(* Logix 5000 project; controller PLC_MCC1201_220AP1 vendor 1 type 14 code 164 rev 35.11; software revision 35.00; part 4 of 25 *)

        [201]   // Flaw Tail Lane Ptr
        [202]   // Flaw Tail Offset Ptr
        [203]   // Count at Sync Pulse to Host MSW
        [204]   // Count at Sync Pulse to Host LSW
        [205]   // Count at Data Request to Host MSW
        [206]   // Count at Data Request to Host LSW
        [207]   // Host Integer location for the number of 1 Meter Pulses(0-39)
        [208]   // Host location for 1/10 millimeter position since last 1 Meter
        [209].0   // Data Request to Host
        [209].1   // Cover Closed to Host
        [209].2   // Use Insp. Booth P.B. only, to host
        [209].4   // Cross Break in Progress to Host
        [209].6   // Image Automation in Alarm to Host
        [209].7   // Image Automation Watchdog Alarm to Host
        [210]   // Lehr Speed to Host
        [211]   // Manual Inspection Flaw Pos. MSW
        [212]   // Manual Inspection Flaw Pos. LSW
        [234]   // Time for last Meter in 0.01 sec
        [237]   // Copy of Count at Data Request to Host MSW
        [238]   // Copy of Count at Data Request to Host LSW
        [209].5   // Crush All Plates to Host
        [209].8   // Always True Signal to Host
   N44 : DINT[213] := ([0] := -1, [2] := -1, [4] := -1, [6] := -1, [8] := -1, [10] := -1, [12] := -1, [14] := -1, [16] := -1, [18] := -1, [20] := -1, [22] := -1, [24] := -1, [26] := -1, [28] := -1, [30] := -1, [32] := -1, [34] := -1, [36] := -1, [38] := -1, [40] := -1, [42] := -1, [44] := -1, [46] := -1, [48] := -1, [50] := -1, [52] := -1, [54] := -1, [56] := -1, [58] := -1, [60] := -1, [62] := -1, [64] := -1, [66] := -1, [68] := -1, [70] := -1, [72] := -1, [74] := -1, [76] := -1, [78] := -1, [80] := -1, [82] := -1, [84] := -1, [86] := -1, [88] := -1, [90] := -1, [92] := -1, [94] := -1, [96] := -1, [98] := -1, [200] := -1);
   N45 : DINT[58] := ([4] := 244, [5] := 129, [6] := 810, [21] := -21856, [23] := 1296, [24] := 253, [26] := 8192, [27] := 5376, [29] := 20480, [30] := 8192, [31] := 8192, [32] := 8192, [33] := 8192, [34] := 8192, [35] := 8192, [36] := 8192, [37] := 8192, [38] := 8192, [39] := 8192, [40] := 8192, [41] := 8192);
   N46 : DINT[7] := ([0] := 142);
        [0]   // Strain Count
        [1]   // Strain Status
        [2]   // Start Strain Cycle
        [3]   // Bar Disable For Reliance
   N47 : DINT[200] := ([0] := 296, [1] := 523, [2] := 448, [3] := 301, [4] := 248, [5] := 289, [6] := 298, [7] := 292, [8] := 287, [9] := 256, [10] := 239, [11] := 185, [12] := 175, [13] := 141, [14] := 116, [15] := 67, [16] := 50, [17] := 74, [18] := 73, [19] := 79, [20] := 75, [21] := 92, [22] := 90, [23] := 90, [24] := 73, [25] := 47, [26] := 29, [27] := 1, [28] := 36, [29] := 39, [30] := 45, [31] := 76, [32] := 75, [33] := 92, [34] := 73, [35] := 84, [36] := 96, [37] := 90, [38] := 74, [39] := 56, [40] := 68, [41] := 72, [42] := 71, [43] := 81, [44] := 78, [45] := 86, [46] := 85, [47] := 88, [48] := 96, [49] := 76, [50] := 54, [51] := 39, [52] := 68, [53] := 89, [54] := 93, [55] := 100, [56] := 103, [57] := 111, [58] := 100, [59] := 114,
        [60] := 125, [61] := 115, [62] := 111, [63] := 109, [64] := 102, [65] := 135, [66] := 135, [67] := 131, [68] := 153, [69] := 136, [70] := 126, [71] := 125, [72] := 122, [73] := 100, [74] := 84, [75] := 82, [76] := 111, [77] := 126, [78] := 127, [79] := 115, [80] := 128, [81] := 123, [82] := 138, [83] := 123, [84] := 110, [85] := 83, [86] := 62, [87] := 68, [88] := 91, [89] := 82, [90] := 100, [91] := 129, [92] := 129, [93] := 110, [94] := 118, [95] := 103, [96] := 121, [97] := 96, [98] := 94, [99] := 107, [100] := 129, [101] := 119, [102] := 123, [103] := 123, [104] := 95, [105] := 101, [106] := 90, [107] := 82, [108] := 78, [109] := 39, [110] := 37, [111] := 62, [112] := 77, [113] := 64, [114] := 68, [115] := 81, [116] := 94, [117] := 83, [118] := 94, [119] := 109,
        [120] := 118, [121] := 123, [122] := 132, [123] := 160, [124] := 190, [125] := 245, [126] := 254, [127] := 295, [128] := 313, [129] := 349, [130] := 383, [131] := 378, [132] := 331, [133] := 284, [134] := 363, [135] := 508, [136] := 87, [137] := 124, [138] := 115, [139] := 132, [140] := 122, [141] := 121, [142] := 126, [143] := 184, [144] := 171, [145] := 122, [146] := 134, [147] := 224, [148] := 143, [149] := 179, [150] := 182, [151] := 488, [152] := 583, [153] := 710, [154] := 493, [155] := 464, [156] := 456, [157] := 470, [158] := 458, [159] := 453, [160] := 458, [161] := 459, [162] := 459, [163] := 464, [164] := 470, [165] := 437, [166] := 467, [167] := 455, [168] := 446, [169] := 426, [170] := 443, [171] := 429, [172] := 422, [173] := 436, [174] := 449, [175] := 433, [176] := 452, [177] := 425, [178] := 447, [179] := 437,
        [180] := 443, [181] := 420, [182] := 440, [183] := 439, [184] := 417, [185] := 427, [186] := 428, [187] := 431, [188] := 429, [189] := 437, [190] := 437, [191] := 419, [192] := 435, [193] := 420, [194] := 421, [195] := 427, [196] := 430, [197] := 439, [198] := 423, [199] := 451);
   N48 : DINT[200] := ([0] := 1032, [1] := 1100, [2] := 1101, [3] := 1081, [4] := 1082, [5] := 1097, [6] := 1100, [7] := 1108, [8] := 1119, [9] := 1115, [10] := 1120, [11] := 1115, [12] := 1114, [13] := 1110, [14] := 1106, [15] := 1095, [16] := 1102, [17] := 1112, [18] := 1121, [19] := 1118, [20] := 1123, [21] := 1120, [22] := 1119, [23] := 1114, [24] := 1118, [25] := 1115, [26] := 1111, [27] := 1106, [28] := 1114, [29] := 1120, [30] := 1125, [31] := 1129, [32] := 1126, [33] := 1119, [34] := 1118, [35] := 1126, [36] := 1126, [37] := 1126, [38] := 1117, [39] := 1117, [40] := 1118, [41] := 1124, [42] := 1124, [43] := 1125, [44] := 1124, [45] := 1128, [46] := 1128, [47] := 1130, [48] := 1132, [49] := 1124, [50] := 1114, [51] := 1115, [52] := 1124, [53] := 1136, [54] := 1133, [55] := 1132, [56] := 1133, [57] := 1133, [58] := 1137, [59] := 1140,
        [60] := 1136, [61] := 1129, [62] := 1125, [63] := 1128, [64] := 1126, [65] := 1134, [66] := 1133, [67] := 1136, [68] := 1139, [69] := 1131, [70] := 1132, [71] := 1140, [72] := 1129, [73] := 1127, [74] := 1115, [75] := 1131, [76] := 1133, [77] := 1135, [78] := 1132, [79] := 1138, [80] := 1140, [81] := 1136, [82] := 1140, [83] := 1138, [84] := 1132, [85] := 1123, [86] := 1128, [87] := 1127, [88] := 1137, [89] := 1133, [90] := 1134, [91] := 1135, [92] := 1132, [93] := 1127, [94] := 1131, [95] := 1129, [96] := 1126, [97] := 1117, [98] := 1120, [99] := 1134, [100] := 1129, [101] := 1130, [102] := 1130, [103] := 1121, [104] := 1119, [105] := 1115, [106] := 1115, [107] := 1116, [108] := 1105, [109] := 1098, [110] := 1102, [111] := 1116, [112] := 1113, [113] := 1108, [114] := 1108, [115] := 1108, [116] := 1113, [117] := 1108, [118] := 1108, [119] := 1107,
        [120] := 1097, [121] := 1094, [122] := 1097, [123] := 1094, [124] := 1092, [125] := 1091, [126] := 1093, [127] := 1089, [128] := 1084, [129] := 1091, [130] := 1089, [131] := 1082, [132] := 1065, [133] := 1068, [134] := 1099, [135] := 1083, [136] := 838, [137] := 839, [138] := 830, [139] := 832, [140] := 829, [141] := 828, [142] := 829, [143] := 827, [144] := 827, [145] := 850, [146] := 846, [147] := 842, [148] := 848, [149] := 846, [150] := 870, [151] := 1103, [152] := 1068, [153] := 1082, [154] := 1031, [155] := 1033, [156] := 1029, [157] := 1034, [158] := 1034, [159] := 1033, [160] := 1035, [161] := 1039, [162] := 1040, [163] := 1038, [164] := 1041, [165] := 1045, [166] := 1041, [167] := 1040, [168] := 1042, [169] := 1041, [170] := 1044, [171] := 1045, [172] := 1040, [173] := 1042, [174] := 1045, [175] := 1040, [176] := 1042, [177] := 1032, [178] := 1041, [179] := 1049,
        [180] := 1042, [181] := 1046, [182] := 1045, [183] := 1043, [184] := 1044, [185] := 1048, [186] := 1047, [187] := 1043, [188] := 1048, [189] := 1040, [190] := 1040, [191] := 1043, [192] := 1041, [193] := 1038, [194] := 1041, [195] := 1042, [196] := 1039, [197] := 1044, [198] := 1038, [199] := 1042);
   N50 : DINT[40] := ([5] := 6278, [7] := 1);
        [39].0   // NO1 CRUSHER Crusher is up and in manual alarm horn has been acknowledged.
   N500 : DINT[24] := ([1] := 1755, [2] := 1755, [3] := 1755, [4] := 1755, [5] := 1755, [6] := 1755, [7] := 1755);
   N501 : DINT[25] := ([1] := 21, [2] := 21, [3] := 21, [4] := 21, [5] := 71, [6] := 71, [7] := 6);
   N502 : DINT[25] := ([1] := 361, [2] := 361, [3] := 361, [4] := 361, [5] := 361, [6] := 361, [7] := 361);
   N504 : DINT[25] := ([1] := 2975, [2] := 2975, [3] := 2975, [4] := 2975, [5] := 3600, [6] := 3600, [7] := 4398);
   N505 : DINT[25] := ([1] := 4229, [2] := 4229, [3] := 4229, [4] := 4229, [5] := 1514, [6] := 1514, [7] := 21881);
   N506 : DINT[25];
   N507 : DINT[25] := ([1] := 765, [2] := 765, [3] := 766, [4] := 766, [5] := 1493, [6] := 1493, [7] := 103, [17] := 1816, [18] := 1816, [24] := 2750);
        [17]   // SPEED CALC Current Command freq. For washer Sponges
        [24]   // SPEED CALC Current Lehr spd + 1.5% Times 10
   N53 : DINT[10];
        [0]   // Disable Y-cuts Information Written FROM Host computer
        [1]   // MANUAL INSPCTN Reject flaw Q.A. Flaw Lamps host Write word
        [2].3   // HOST WRITE Inhibit bit For Trim Deck E-stop
        [2].4   // HOST WRITE Inhibit bit For Critical Failure
        [2].5   // HOST WRITE Inhibit bit For trim Deck drive Fault
        [2].7   // HOST WRITE Inhibit bit for Mainline Backup
        [2].8   // HOST WRITE Inhibit bit for Drive system E-stop
        [2].10   // HOST WRITE Inhibit bit for Sec. Trans. Drive fault
        [2].11   // Host Critical Alarm Present
        [2].12   // View TEC15V alarm present
        [2].13   // APC Low Alarm
        [3].0   // From Host Enable 37B's REV controls
        [5].0   // ISRA 5D System QC Request Signal
        [5].1   // ISRA 5D System Cut Signal
        [8].6   // Z200 Reset Alarms
        [8]   // HOST WRITE DATA: ZONE 200 (Cutting Area) HMI Commands
        [8].0   // Z200 Start Cycle
        [8].3   // Z200 Stop Cleaning
        [8].1   // Z200 Stop Cycle
        [8].4   // Z200 Zone in Automatic
        [8].5   // Z200 Zone in Manual
        [8].2   // Z200 Start Cleaning
        [7]   // HOST WRITE DATA: ZONE UPS (Drop Conveyor Area) HMI Commands
        [7].0   // ZUPS Start Cycle
        [7].1   // ZUPS Stop Cycle
        [7].2   // ZUPS Start Cleaning
        [7].3   // ZUPS Stop Cleaning
        [7].4   // ZUPS Zone in Automatic
        [7].5   // ZUPS Zone in Manual
        [7].6   // ZUPS Reset Alarms
   N53_HOST : INT[10];
   N54 : DINT[501] := ([200] := 516, [201] := 1844, [202] := 516, [203] := 516, [204] := 516, [206] := 4, [207] := 31, [208] := 514, [211] := 176, [239] := 16, [240] := -65524, [244] := 4096, [246] := 512, [247] := 256, [248] := 512, [249] := 1, [250] := 15, [251] := 17, [252] := 12, [253] := 8, [254] := 44, [255] := 27, [256] := 15, [257] := 13, [258] := 10, [259] := 10, [260] := 481, [261] := 480, [262] := 481, [264] := -32287, [265] := 10, [266] := 110, [270] := 132, [271] := 164, [273] := 1, [274] := 1, [275] := 1, [276] := 1, [277] := 1, [281] := -32768, [341] := 133, [368] := -11667, [410] := 9, [411] := 510, [420] := 6234);
        [200].1   // RIBBON WASHER BRUSH #1 AUTO Mode Bit
        [200].2   // RIBBON WASHER BRUSH #1 MANUAL Mode Bit
        [200].3   // RIBBON WASHER BRUSH #1 ON Sw. Inputs
        [200].4   // RIBBON WASHER BRUSH #1 OFF Sw. Inputs
        [200].5   // RIBBON WASHER BRUSH #1 UPPER RETRACT Sw. Inputs
        [200].6   // RIBBON WASHER BRUSH #1 UPPER CONVERGE Sw. Inputs
        [200].7   // RIBBON WASHER BRUSH #1 LOWER RETRACT Sw. Inputs
        [200].8   // RIBBON WASHER BRUSH #1 LOWER CONVERGE Sw. Inputs
        [200].9   // RIBBON WASHER BRUSH #1 Manual Mode Lamp
        [200].10   // RIBBON WASHER BRUSH #1 OFF selected Manual mode
        [202].1   // RIBBON WASHER SPONGE UNIT AUTO Mode Bit
        [202].2   // RIBBON WASHER SPONGE UNIT MANUAL Mode Bit
        [202].3   // RIBBON WASHER SPONGE UNIT ON Sw. Inputs
        [202].4   // RIBBON WASHER SPONGE UNIT OFF Sw. Inputs
        [202].5   // RIBBON WASHER SPONGE UNIT UPPER RETRACT Sw. Inputs
        [202].6   // RIBBON WASHER SPONGE UNIT UPPER CONVERGE Sw. Inputs
        [202].7   // RIBBON WASHER SPONGE UNIT LOWER RETRACT Sw. Inputs
        [202].8   // RIBBON WASHER SPONGE UNIT LOWER CONVERGE Sw. Inputs
        [202].9   // RIBBON WASHER SPONGE UNIT Manual Mode Lamp
        [202].10   // RIBBON WASHER SPONGE UNIT OFF selected Manual mode
        [203].1   // RIBBON WASHER AIR KNIFE AUTO Mode Bit
        [203].2   // RIBBON WASHER AIR KNIFE MANUAL Mode Bit
        [203].3   // RIBBON WASHER AIR KNIFE UNIT #1 RETRACT Sw. Inputs
        [203].4   // RIBBON WASHER AIR KNIFE UNIT #1 CONVERGE Sw. Inputs
        [203].5   // RIBBON WASHER AIR KNIFE UNIT #2 RETRACT Sw. Inputs
        [203].6   // RIBBON WASHER AIR KNIFE UNIT #2 CONVERGE Sw. Inputs
        [203].7   // RIBBON WASHER AIR KNIFE BLOWER ON WASH-AK-ON
        [203].8   // RIBBON WASHER AIR KNIFE BLOWER OFF WASH-AK-OFF
        [203].9   // RIBBON WASHER AIR KNIFE Manual Mode Lamp
        [203].10   // RIBBON WASHER AIR KNIFE BLOWER MANUAL OFF WASH-AK-MOFF
        [204].1   // RIBBON WASHER WATER SPRAYERS AUTO Mode Bit
        [204].2   // RIBBON WASHER WATER SPRAYERS MANUAL Mode Bit
        [204].3   // RIBBON WASHER WATER SPRAYERS ON Sw. Inputs
        [204].4   // RIBBON WASHER WATER SPRAYERS OFF Sw. Inputs
        [204].5   // RIBBON WASHER WATER SPRAYERS
        [204].6   // RIBBON WASHER WATER SPRAYERS
        [204].7   // RIBBON WASHER WATER SPRAYERS
        [204].8   // RIBBON WASHER WATER SPRAYERS
        [204].9   // RIBBON WASHER WATER SPRAYERS Manual Mode Lamp
        [205].1   // RIBBON WASHER BRUSH #1 UPPER CONVERGE Output
        [205].3   // RIBBON WASHER SPONGE UPPER CONVERGE Output
        [205].4   // RIBBON WASHER AIR KNIFE #1 UPPER CONVERGE Output
        [205].5   // RIBBON WASHER AIR KNIFE #2 UPPER CONVERGE Output
        [205].6   // RIBBON WASHER BRUSH #1 Water valve Output
        [205].7   // RIBBON WASHER BRUSH #2 Water valve Output
        [205].8   // RIBBON WASHER SPONGE Water valve Output
        [205].9   // RIBBON WASHER Master Water valve Output
        [206].1   // RIBBON WASHER BRUSH #1 LOWER CONVERGE Output
        [206].3   // RIBBON WASHER SPONGE LOWER CONVERGE Output
        [206].4   // RIBBON WASHER AIR KNIFE #1 LOWER CONVERGE Output
        [206].5   // RIBBON WASHER AIR KNIFE #2 LOWER CONVERGE Output
        [207].0   // RIBBON WASHER Crossbreak Acknowledge 0 = Ack'd 1 = Must Ack
        [207].1   // RIBBON WASHER BRUSH #1 Crossbreak Active
        [207].2   // RIBBON WASHER BRUSH #2 Crossbreak Active
        [207].3   // RIBBON WASHER SPONGE Crossbreak Active
        [207].4   // RIBBON WASHER AIR KNIFE #1 Crossbreak Active
        [207].5   // RIBBON WASHER AIR KNIFE #2 Crossbreak Active
        [207].6   // Water Spray Solenoid #3 Crossbreak Active
        [207].7   // RIBBON WASHER Crossbreak Reset (Two P.B.s ANDed)
        [208].1   // Eclipse Mode On Permissive
        [208].2   // Eclipse Mode Off Permissive
        [208].3   // RIBBON WASHER Ribbon is an Active product (Active mode ON)
        [211].0   // WASHER-BR1 UP Drive Fault - MMI Reporting
        [211].1   // WASHER-BR1 LO Drive Fault - MMI Reporting
        [211].2   // WASHER-BR2 UP Drive Fault - MMI Reporting
        [211].3   // WASHER-BR2 LO Drive Fault - MMI Reporting
        [211].4   // WASHER-SPG UP Drive Fault - MMI Reporting
        [211].5   // WASHER-SPG LO Drive Fault - MMI Reporting
        [212].0   // WASHER-BR1 UP Drive Forward - MMI Reporting
        [212].1   // WASHER-BR1 LO Drive Forward - MMI Reporting
        [212].2   // WASHER-BR2 UP Drive Forward - MMI Reporting
        [212].3   // WASHER-BR2 LO Drive Forward - MMI Reporting
        [212].4   // WASHER-SPG UP Drive Forward - MMI Reporting
        [212].5   // WASHER-SPG LO Drive Forward - MMI Reporting
        [213].0   // WASHER-BR1 UP SS1 - MMI Reporting
        [213].1   // WASHER-BR1 LO SS1 - MMI Reporting
        [213].2   // WASHER-BR2 UP SS1 - MMI Reporting
        [213].3   // WASHER-BR2 LO SS1 - MMI Reporting
        [213].4   // WASHER-SPG UP SS1 - MMI Reporting
        [213].5   // WASHER-SPG LO SS1 - MMI Reporting
        [213].8   // WASHER-BR1 UP SS2 - MMI Reporting
        [213].9   // WASHER-BR1 LO SS2 - MMI Reporting
        [213].10   // WASHER-BR2 UP SS2 - MMI Reporting
        [213].11   // WASHER-BR2 LO SS2 - MMI Reporting
        [213].12   // WASHER-SPG UP SS2 - MMI Reporting
        [213].13   // WASHER-SPG LO SS2 - MMI Reporting
        [239].0   // NO. 1 CRUSHER Drive Operating Forward bit - MMI Reporting
        [239].2   // NO. 1 CRUSHER SS1 Input Selected - MMI reporting
        [239].4   // NO. 1 CRUSHER SS2 input Selected
        [239].8   // NO. 1 CRUSHER Drive faulted
        [240].0   // NO. 1 CRUSHER Auto drop Prohibited!
        [240].1   // NO. 1 CRUSHER Automatic Mode
        [240].2   // NO. 1 CRUSHER Manual Mode
        [240].3   // NO. 1 CRUSHER Crusher drive E-Stop
        [240].4   // NO. 1 CRUSHER Crusher drive Control system Failure
        [240].5   // No. 1 Crusher Beater bar Drive fault
        [240].6   // NO. 1 CRUSHER Cullet system Failure
        [240].8   // NO. 1 CRUSHER one shot!
        [240].10   // NO. 1 CRUSHER Crusher down In auto mode After Power Loss
        [240].11   // NO. 1 CRUSHER Generator Supplying Power to No. 1 Crusher
        [240].13   // NO. 1 CRUSHER Automatic Drop conditions
        [240].14   // No. 1 CRUSHER Down Proximity Sw.
        [240].15   // NO. 1 CRUSHER Up Proximity sw.
        [241].0   // NO. 1 CRUSHER Control Tech. Drive system E-stop
        [241].1   // NO. 1 CRUSHER Control Tech. Master Drive system Critical fail
        [241].2   // NO. 1 CRUSHER Control Tech. Drive system Drive fault
        [241].6   // NO. 1 CRUSHER Trim deck Drive system E-stop
        [241].7   // NO. 1 CRUSHER Trim deck Drive system Critical fail
        [241].8   // NO. 1 CRUSHER Trim deck Drive system Drive fault
        [242].0   // NO. 1 CRUSHER Drop Crusher Push-buton Rel. console
        [242].1   // NO. 1 CRUSHER Mainline Backup to Trim deck
        [242].6   // NO. 1 CRUSHER Sec. trans. Drive system E-stop
        [242].8   // NO. 1 CRUSHER Sec. trans. Drive system Drive fault
        [244].0   // NO. 1 CRUSHER Reliance Drive system E-stop INIBIT BIT
        [244].1   // NO. 1 CRUSHER Reliance Drive system Critical fail INIBIT BIT
        [244].2   // NO. 1 CRUSHER Reliance Drive system Drive fault INIBIT BIT
        [244].3   // NO. 1 CRUSHER FUTURE INIBIT BIT
        [244].4   // NO. 1 CRUSHER FUTURE INIBIT BIT
        [244].5   // NO. 1 CRUSHER FUTURE INIBIT BIT
        [244].6   // NO. 1 CRUSHER Trim deck Drive system E-stop INIBIT BIT
        [244].7   // NO. 1 CRUSHER Trim deck Drive system Critical fail INIBIT BIT
        [244].8   // NO. 1 CRUSHER Trim deck Drive system Drive fault INIBIT BIT
        [244].9   // NO. 1 CRUSHER FUTURE INIBIT BIT
        [244].10   // NO. 1 CRUSHER FUTURE INIBIT BIT
        [244].11   // NO. 1 CRUSHER FUTURE INIBIT BIT
        [244].12   // NO. 1 CRUSHER FUTURE INIBIT BIT
        [244].13   // NO. 1 CRUSHER FUTURE INIBIT BIT
        [244].14   // NO. 1 CRUSHER FUTURE INIBIT BIT
        [244].15   // NO. 1 CRUSHER FUTURE INIBIT BIT
        [245].1   // NO. 1 CRUSHER Mainline Backup to Trim deck INIBIT BIT
        [245].6   // NO. 1 CRUSHER Sec. trans. Drive system E-stop INIBIT BIT
        [245].7   // NO. 1 CRUSHER Sec. trans. Drive system Critical fail INIBIT BIT
        [245].8   // NO. 1 CRUSHER Sec. trans. Drive system Drive fault INIBIT BIT
        [246]   // NO.1 CRUSHER Drop reason History stack Word 1 of 3
        [246].0   // NO. 1 CRUSHER Reliance Drive system E-stop HISTORY BIT
        [246].1   // NO. 1 CRUSHER Reliance Drive system Critical fail HISTORY BIT
        [246].2   // NO. 1 CRUSHER Reliance Drive system Drive fault HISTORY BIT
        [246].3   // NO. 1 CRUSHER SPARE HISTORY BIT
        [246].4   // NO. 1 CRUSHER Trim deck Drive system E-stop HISTORY BIT
        [246].5   // NO. 1 CRUSHER Trim deck Drive system Critical fail HISTORY BIT
        [246].6   // NO. 1 CRUSHER Trim deck Drive system Drive fault HISTORY BIT
        [246].7   // NO. 1 CRUSHER SPARE HISTORY BIT
        [246].8   // NO. 1 CRUSHER Drop crusher Pushbutton HISTORY BIT
        [246].9   // NO. 1 CRUSHER Mainlin backup HISTORY BIT
        [246].10   // NO. 1 CRUSHER SPARE HISTORY BIT
        [246].11   // NO. 1 CRUSHER SPARE HISTORY BIT
        [246].12   // NO. 1 CRUSHER Sec. Trans. Drive system E-stop HISTORY BIT
        [246].13   // NO. 1 CRUSHER Sec. Trans. Drive system Critical fail HISTORY BIT
        [246].14   // NO. 1 CRUSHER Sec. Trans. Drive system Drive fault HISTORY BIT
        [246].15   // NO. 1 CRUSHER Power-loss Failure HISTORY BIT
        [247]   // NO. 1 CRUSHER Drop reason Hirtory stack Word 2 of 3
        [247].0   // NO. 1 CRUSHER FUTURE
        [247].1   // NO. 1 CRUSHER FUTURE
        [247].2   // NO. 1 CRUSHER FUTURE
        [247].3   // NO. 1 CRUSHER FUTURE
        [247].4   // NO. 1 CRUSHER FUTURE
        [247].5   // NO. 1 CRUSHER FUTURE
        [247].6   // NO. 1 CRUSHER FUTURE
        [247].7   // NO. 1 CRUSHER FUTURE
        [247].8   // NO. 1 CRUSHER FUTURE
        [247].9   // NO. 1 CRUSHER FUTURE
        [247].10   // NO. 1 CRUSHER FUTURE
        [247].11   // NO. 1 CRUSHER FUTURE
        [247].12   // NO. 1 CRUSHER FUTURE
        [247].13   // NO. 1 CRUSHER FUTURE
        [247].14   // NO. 1 CRUSHER FUTURE
        [247].15   // NO. 1 CRUSHER FUTURE
        [248]   // NO.1 CRUSHER Drop reason History stack Word 3 of 3
        [248].0   // NO. 1 CRUSHER FUTURE
        [248].1   // NO. 1 CRUSHER FUTURE
        [248].2   // NO. 1 CRUSHER FUTURE
        [248].3   // NO. 1 CRUSHER FUTURE
        [248].4   // NO. 1 CRUSHER FUTURE
        [248].5   // NO. 1 CRUSHER FUTURE
        [248].6   // NO. 1 CRUSHER FUTURE
        [248].7   // NO. 1 CRUSHER FUTURE
        [248].8   // NO. 1 CRUSHER FUTURE
        [248].9   // NO. 1 CRUSHER FUTURE
        [248].10   // NO. 1 CRUSHER FUTURE
        [248].11   // NO. 1 CRUSHER FUTURE
        [248].12   // NO. 1 CRUSHER FUTURE
        [248].13   // NO. 1 CRUSHER FUTURE
        [248].14   // NO. 1 CRUSHER FUTURE
        [248].15   // NO. 1 CRUSHER FUTURE
        [249]   // NO. 1 CRUSHER Drop reason History stack Time Word (Hour) 1 of 3
        [250]   // NO. 1 CRUSHER Drop reason History stack Time Word (Hour) 2 of 3
        [251]   // NO. 1 CRUSHER Drop reason History stack Time Word (Hour) 3 of 3
        [252]   // NO. 1 CRUSHER Drop reason History stack Time Word (Min) 1 of 3
        [253]   // NO. 1 CRUSHER Drop reason History stack Time Word (Min) 2 of 3
        [254]   // NO. 1 CRUSHER Drop reason History stack Time Word (Min) 3 of 3
        [255]   // NO. 1 CRUSHER Drop reason History stack Month Word 1 of 3
        [256]   // NO. 1 CRUSHER Drop reason History stack Month Word 2 of 3
        [257]   // NO. 1 CRUSHER Drop reason History stack Month Word 3 of 3
        [258]   // NO. 1 CRUSHER Drop reason History stack Day Word 1 of 3
        [259]   // NO. 1 CRUSHER Drop reason History stack Day Word 2 of 3
        [260].0   // CRSSBRK ZONE 1 Crossbreak In progress Lamp * INSIDE LEHR *
        [260].1   // CRSSBRK ZONE 1 North Outside Bypass Switch ON=Bypass OFF=Operate
        [260].2   // CRSSBRK ZONE 1 North Inside Bypass Switch ON=Bypass OFF=Operate
        [260].3   // CRSSBRK ZONE 1 South Outside Bypass Switch ON=Bypass OFF=Operate
        [260].4   // CRSSBRK ZONE 1 South Inside Bypass Switch ON=Bypass OFF=Operate
        [260].5   // CRSSBRK ZONE 1 North Outside Photo-eye ALARM WHEN P.E. IS CLEAR
        [260].6   // CRSSBRK ZONE 1 North Inside Photo-eye ALARM WHEN P.E. IS CLEAR
        [260].7   // CRSSBRK ZONE 1 South Outside Photo-eye ALARM WHEN P.E. IS CLEAR
        [260].8   // CRSSBRK ZONE 1 South Inside Photo-eye ALARM WHEN P.E. IS CLEAR
        [260].9   // CRSSBRK ZONE 1 North Outside Lamp ON=Bypass OFF=Normal
        [260].10   // CRSSBRK ZONE 1 North Inside Lamp ON=Bypass OFF=Normal
        [260].11   // CRSSBRK ZONE 1 South Outside Lamp ON=Bypass OFF=Normal
        [260].12   // CRSSBRK ZONE 1 South Inside Lamp ON=Bypass OFF=Normal
        [260].14   // CRSSBRK ZONE 1 Crossbreak has Been Acknowledged
        [260].15   // CRSSBRK ZONE 1 Alarm horn Silence One shot
        [261].0   // CRSSBRK ZONE 2 Crossbreak In progress Lamp * LEHR EXIT *
        [261].1   // CRSSBRK ZONE 2 North Outside Bypass Switch ON=Bypass OFF=Operate
        [261].2   // CRSSBRK ZONE 2 North Inside Bypass Switch ON=Bypass OFF=Operate
        [261].3   // CRSSBRK ZONE 2 South Outside Bypass Switch ON=Bypass OFF=Operate
        [261].4   // CRSSBRK ZONE 2 South Inside Bypass Switch ON=Bypass OFF=Operate
        [261].5   // CRSSBRK ZONE 2 North Outside Photo-eye ALARM WHEN P.E. IS CLEAR
        [261].6   // CRSSBRK ZONE 2 North Inside Photo-eye ALARM WHEN P.E. IS CLEAR
        [261].7   // CRSSBRK ZONE 2 South Outside Photo-eye ALARM WHEN P.E. IS CLEAR
        [261].8   // CRSSBRK ZONE 2 South Inside Photo-eye ALARM WHEN P.E. IS CLEAR
        [261].9   // CRSSBRK ZONE 2 North Outside Lamp ON=Bypass OFF=Normal
        [261].10   // CRSSBRK ZONE 2 North Inside Lamp ON=Bypass OFF=Normal
        [261].11   // CRSSBRK ZONE 2 South Outside Lamp ON=Bypass OFF=Normal
        [261].12   // CRSSBRK ZONE 2 South Inside Lamp ON=Bypass OFF=Normal
        [262].0   // CRSSBRK ZONE 3 Crossbreak In progress Lamp * RIBBON WASHER
        [262].1   // CRSSBRK ZONE 3 North Outside Bypass Switch ON=Bypass OFF=Operate
        [262].2   // CRSSBRK ZONE 3 North Inside Bypass Switch ON=Bypass OFF=Operate
        [262].3   // CRSSBRK ZONE 3 South Outside Bypass Switch ON=Bypass OFF=Operate
        [262].4   // CRSSBRK ZONE 3 South Inside Bypass Switch ON=Bypass OFF=Operate
        [262].5   // CRSSBRK ZONE 3 North Outside Photo-eye ALARM WHEN P.E. IS CLEAR
        [262].6   // CRSSBRK ZONE 3 North Inside Photo-eye ALARM WHEN P.E. IS CLEAR
        [262].7   // CRSSBRK ZONE 3 South Outside Photo-eye ALARM WHEN P.E. IS CLEAR
        [262].8   // CRSSBRK ZONE 3 South Inside Photo-eye ALARM WHEN P.E. IS CLEAR
        [262].9   // CRSSBRK ZONE 3 North Outside Lamp ON=Bypass OFF=Normal
        [262].10   // CRSSBRK ZONE 3 North Inside Lamp ON=Bypass OFF=Normal
        [262].11   // CRSSBRK ZONE 3 South Outside Lamp ON=Bypass OFF=Normal
        [262].12   // CRSSBRK ZONE 3 South Inside Lamp ON=Bypass OFF=Normal
        [263].1   // CRSSBRK ZONE 4 North Outside Bypass Switch ON=Bypass OFF=Operate
        [263].5   // CRSSBRK ZONE 4 North Outside Photo-eye ALARM WHEN P.E. IS CLEAR
        [263].14   // FIX MMI IAL TEMPERATURE ALARM
        [264].0   // CRSSBRK ZONE 5 Crossbreak In progress Lamp * MAN INSPCT *
        [264].1   // CRSSBRK ZONE 5 North Outside Bypass Switch ON=Bypass OFF=Operate
        [264].2   // CRSSBRK ZONE 5 North Inside Bypass Switch ON=Bypass OFF=Operate
        [264].3   // CRSSBRK ZONE 5 South Outside Bypass Switch ON=Bypass OFF=Operate
        [264].4   // CRSSBRK ZONE 5 South Inside Bypass Switch ON=Bypass OFF=Operate
        [264].5   // CRSSBRK ZONE 5 North Outside Photo-eye ALARM WHEN P.E. IS CLEAR
        [264].6   // CRSSBRK ZONE 5 North Inside Photo-eye ALARM WHEN P.E. IS CLEAR
        [264].7   // CRSSBRK ZONE 5 South Outside Photo-eye ALARM WHEN P.E. IS CLEAR
        [264].8   // CRSSBRK ZONE 5 South Inside Photo-eye ALARM WHEN P.E. IS CLEAR
        [264].9   // CRSSBRK ZONE 5 North Outside Lamp ON=Bypass OFF=Normal
        [264].10   // CRSSBRK ZONE 5 North Inside Lamp ON=Bypass OFF=Normal
        [264].11   // CRSSBRK ZONE 5 South Outside Lamp ON=Bypass OFF=Normal
        [264].12   // CRSSBRK ZONE 5 South Inside Lamp ON=Bypass OFF=Normal
        [264].15   // MARKING BRIDGE Cross break Present At Marking Bridge
        [265]   // NO. 1 CRUSHER Drop reason History stack Day Word 3 of 3
        [266]   // APC Lehr Speed Multiplier
        [267].0   // ISRA 5D 24VDC OK
        [267].1   // ISRA 5D System Watchdog
        [267].2   // ISRA 5D 12V DC OK
        [267].3   // ISRA 5D System Ok
        [267].4   // ISRA 5D System Warning
        [267].5   // ISRA 5D System Error 1
        [267].6   // ISRA 5D System Error 2
        [267].7   // ISRA 5D Crossbreak at 5D
        [281].5   // IMAGE AUTO Retro cover Closed
        [281].6   // IMAGE AUTO Retro cover Closure alrm Acknowledge
        [281].7   // IMAGE AUTO Retro cover Closure Alarm
        [281].11   // one shot!
        [282]   // Storage for Crossbreak Tracking to IAL
        [291].0   // MANUAL INSPCTN Booth Flaw Push-Button
        [291].1   // MANUAL INSPCTN Booth Reject Push-Button
        [292].9   // HOST READ DATA: Low-e Inpsection Pulse Entire Ribbon Button
        [292].11   // HOST READ DATA: Low-e Inpsection Spray Right Edge of Ribbon
        [292].12   // HOST READ DATA: Low-e Inpsection Spray Right-Center Lane of Ribbon
        [292].13   // HOST READ DATA: Low-e Inpsection Spray Center Lane of Ribbon
        [292].14   // HOST READ DATA: Low-e Inpsection Spray Left-Center Lane of Ribbon
        [292].15   // HOST READ DATA: Low-e Inpsection Spray Left Edge of Ribbon
        [301].0   // Reliance Data Request Bit
        [301].1   // Reliance Two inch Lehe Pulse
        [341]   // Top Sheet Temperature [0-300 degF]
        [351].0   // TO Host APC Off
        [351].2   // APC low Alarm
        [372].0   // Vibrating Pan Mapped Speed For MMI Read VP917067
        [372].3   // Vibrating Pan Mapped Speed For MMI Read VP917066
        [372].6   // Vibrating Pan Mapped Speed For MMI Read VP917065
        [372].9   // Vibrating Pan Mapped Speed For MMI Read VP917070
        [372].12   // Vibrating Pan Mapped Speed For MMI Read VP917071
        [372].15   // Vibrating Pan Mapped Speed For MMI Read VP917077
        [373].2   // MMI READ Cullet System M32 Sleep Mode Enabled
        [373].3   // MMI READ Cullet System M33 Sleep Mode Enabled
        [373].6   // Vibrating Pan Mapped Speed For MMI Read VP917076
        [373].9   // Vibrating Pan Mapped Speed For MMI Read VP917075
        [373].12   // Vibrating Pan Mapped Speed For MMI Read VP917074
        [373].15   // Vibrating Pan Mapped Speed For MMI Read VP917073
        [374].2   // Vibrating Pan Mapped Speed For MMI Read VP917068
        [374].7   // Vibrating Pan Mapped Speed For MMI Read VP917069
        [374].12   // Vibrating Pan Mapped Speed For MMI Read VP917072
        [374].15   // Vibrating Pan Mapped Speed for MMI Read VP917060
        [375].14   // MMI Read Cullet System M43 Sleep Mode Enabled
        [375].15   // MMI Read Cullet System M41 Sleep Mode Enabled
        [376].0   // MMI Read Cullet System M42 Sleep Mode Enabled
        [376].1   // MMI Read Cullet System M40 Sleep Mode Enabled
        [376].8   // MMI Read Cullet System VP917071 Sleep Mode Enabled
        [376].9   // MMI Read Cullet System VP917070 Sleep Mode Enabled
        [410]   // 0.1mm Pulses Captured on 1 Meter of Travel MSD
        [411]   // 0.1mm Pulses Captured on 1 Meter of Travel LSD
        [420]   // Glass Travel Pulse Count (Counts 50mm Pulses reset @ 10000)
        [301].3   // CRUSH ALL PLATES
        [270]   // ZONE 200 (CUTTING AREA) HMI FEEDBACKS
        [270].7   // Z200 Alarm Presence
        [270].0   // Z200 Cycle Starting
        [270].2   // Z200 Cycle in Stop
        [270].3   // Z200 Cleaning Request
        [270].4   // Z200 Cleaning ON
        [273]   // M203 Drop Conveyor Mode (1 = Down, 2 = Up, 4 = Req Down, 8 = Req Up)
        [270].1   // Z200 Cycle ON
        [270].5   // Z200 in Manual
        [270].6   // Z200 in Automatic
        [274]   // M203 Drop Conveyor Status (1 = Idle, 3 = Moving up/down, 7 = Anomaly)
        [275]   // M205 Breaker Status (1 = Idle, 3 = Running, 7 = Anomaly)
        [276]   // M225 Emergency Xcut Flyer Mode (1 = Manual, 4 = Automatic, 7 = Semiauto)
        [277]   // M225 Emergency Xcut Flyer Status (1 = Idle, 3 =Running, 7 = Anomaly)
        [271]   // ZONE UPS (DROP CONVEYOR AREA) HMI FEEDBACKS
        [271].0   // ZUPS Cycle Starting
        [271].1   // ZUPS Cycle ON
        [271].2   // ZUPS Cycle in Stop
        [271].3   // ZUPS Cleaning Request
        [271].4   // ZUPS Cleaning ON
        [271].5   // ZUPS in Manual
        [271].6   // ZUPS in Automatic
        [271].7   // ZUPS Alarm Presence
   N541 : ALIAS FOR N54[420];
   N54_HOST : INT[501] := ([200] := 516, [201] := 1844, [202] := 516, [203] := 516, [204] := 516, [206] := 4, [207] := 31, [208] := 514, [211] := 176, [239] := 16, [240] := 12, [244] := 4096, [246] := 512, [247] := 256, [248] := 512, [249] := 1, [250] := 15, [251] := 17, [252] := 12, [253] := 8, [254] := 44, [255] := 27, [256] := 15, [257] := 13, [258] := 10, [259] := 10, [260] := 481, [261] := 480, [262] := 481, [264] := -32287, [265] := 10, [266] := 110, [270] := 132, [271] := 164, [273] := 1, [274] := 1, [275] := 1, [276] := 1, [277] := 1, [281] := -32768, [341] := 133, [368] := -11667, [410] := 9, [411] := 510, [420] := 6234);
   N55 : DINT[1];
   N60 : DINT[420] := ([1] := 268, [2] := 800, [11] := 448, [12] := 150, [400] := -32765, [401] := 2706, [402] := 2683, [410] := 2683);
        [1]   // Current lehr Speed
        [2]   // Current trim Speed
        [11]   // Milliseconds Required for 2
        [12]   // Milliseconds Required for 2
        [10]   // Speed for cullet system ???
   N61 : DINT[100] := ([1] := 6, [2] := 254, [5] := 580, [30] := 112, [53] := 1280, [59] := 4095, [61] := 4095, [63] := 4095, [65] := 4095, [67] := 4095, [69] := 4095, [71] := 4095);
        [0].0   // Write New Configuration to Washer Panel Analog Input (Manually set to 1)
        [1]   // VMCC-W1 Analog Input Card Read Data:
        [1].0   // VMCC-W1 Analog Input Card Read Data: Power Up Bit
        [5]   // Top Sheet Temperature Value in Raw units
   N7 : DINT[250] := ([0] := 980, [1] := 532, [2] := 345, [3] := 930, [4] := 1687, [5] := 1, [8] := 2, [9] := 1, [10] := 8, [11] := 3020, [12] := 3028, [13] := 8, [14] := 2970, [15] := 2978, [16] := 1763, [17] := 76, [18] := 12, [19] := 1450, [20] := -1, [21] := 930, [22] := 6899, [23] := 32767, [24] := 32767, [31] := 1081, [32] := 101, [33] := 1031, [34] := 44, [35] := 25602, [36] := 4096, [37] := 1024, [41] := 1337, [42] := 12, [43] := 1031, [44] := 43, [45] := -14078, [46] := 8192, [47] := 1024, [60] := 3072, [161] := 4088, [162] := 4095, [168] := 4095, [171] := 2048, [180] := -1, [181] := -1, [182] := 1, [183] := 1, [201] := 80, [202] := 10, [203] := 1031, [205] := 2, [240] := 20);
        [0]   // Output Index (Gun Bridge)
        [1]   // Distance (cm) From Gun Bridge to Hand Off
        [2]   // Current Sync Pulse Value (cm)
        [3]   // Next Sync Pulse Count Value (cm)
        [4]   // Flaw Position in Track File
        [5]   // Flaw Lane To Output Image Trans. Table 2nd Index
        [6]   // Flaw Lane To Output Image Trans. Table Index
        [7]   // Scanner Number" minus 1 (0 - 4)
        [7].0   // Scanner Number is Odd
        [8]   // FOR Loop Counter For Spray Length
        [9]   // FOR Lpop Counter For Flaw Queue Process
        [10]   // Current Count LSD/100
        [11]   // Current Count MSD*10 (1000/100)
        [12]   // Current Count/100 into One Word (cm)
        [13]   // Sync Count LSD/100
        [14]   // Sync Count MSD*10 (1000/100)
        [15]   // Sync Count /100 into One Word
        [16]   // Start of Gun Test Count (cm)
        [17]   // Gun Test Position (cm) From Start To Current Spray Point
        [18]   // Gun Test Position modulo 16
        [22]   // Number of Skipped Sync Pulses
        [23]   // Time of Longest Read
        [24]   // Longest Delay for New Data
        [30].13   // Host Read Done
   N70 : DINT[3] := ([1] := 59, [2] := 60);
        [1]   // Millisecond Accumulator For 2
   N75 : DINT[2] := ([0] := 800, [1] := 150);
   N80 : DINT[16] := ([0] := 873, [1] := 34);
        [0]   // Time period for last 1 Meter pulse wave
        [1]   // Count of 1Meter pulses from VHSC card(Rollover at 40)
   N9 : DINT[20] := ([0] := 331, [1] := 64, [10] := 980, [15] := 800, [16] := 33);
        [5].1   // Cross Break at Gun Bridge
        [5].2   // I/A Reflector Cover Close
   N98 : DINT[20] := ([0] := -32765, [1] := 2706, [2] := 2683, [4] := 2683, [5] := 2683, [6] := 16, [10] := 414, [11] := 282, [12] := 281, [13] := 269, [14] := 282, [15] := 277);
        [0]   // LEHR SPEED Calculation & Conditioning Status Bits
        [0].0   // LEHR SPEED Speed received From Reliance AutoMax PLC Is Valid
        [0].1   // LEHR SPEED Speed received From Reliance Capping system is Valid
        [0].15   // LEHR SPEED one shot!
        [1]   // LEHR SPEED Value to be Reported to M5 For AutoMax Lehr speed
        [2]   // LEHR SPEED Value to be Reported to M5 For average Lehr speed
        [3]   // LEHR SPEED Value to be Reported to M5 For standard Deviation
        [4]   // LEHR SPEED Value to be Reported to M5 as Reliance Lehr speed
        [5]   // LEHR SPEED Value to be Reported to M5 For current Lehr Speed
        [10]   // DEBUG: Half the Period for 1M pulse at Automax Speed Plus 15IPM [.01 sec]
        [11]   // DEBUG: Lehr Speed from Capping above Automax Speed Plus 15IPM FIFO 1
        [12]   // DEBUG: Lehr Speed from Capping above Automax Speed Plus 15IPM FIFO 2
        [13]   // DEBUG: Lehr Speed from Capping above Automax Speed Plus 15IPM FIFO 3
        [14]   // DEBUG: Lehr Speed from Capping above Automax Speed Plus 15IPM FIFO 4
        [15]   // DEBUG: Lehr Speed from Capping above Automax Speed Plus 15IPM FIFO 5
   N99 : DINT[1000] := ([0] := 2683, [1] := 2683, [2] := 2683, [3] := 2683, [4] := 2683, [5] := 2683, [6] := 2683, [7] := 2683, [8] := 2683, [9] := 2683, [10] := 2683, [11] := 2683, [12] := 2683, [13] := 2683, [14] := 2683, [15] := 2683, [16] := 2683, [17] := 2683, [18] := 2683, [19] := 2683, [20] := 2683, [21] := 2683, [22] := 2683, [23] := 2683, [24] := 2683, [25] := 2683, [26] := 2683, [27] := 2683, [28] := 2683, [29] := 2683, [30] := 2683, [31] := 2683, [32] := 2683, [33] := 2683, [34] := 2683, [35] := 2683, [36] := 2683, [37] := 2683, [38] := 2683, [39] := 2683, [40] := 2683, [41] := 2683, [42] := 2683, [43] := 2683, [44] := 2683, [45] := 2683, [46] := 2683, [47] := 2683, [48] := 2683, [49] := 2683, [50] := 2683, [51] := 2683, [52] := 2683, [53] := 2683, [54] := 2683, [55] := 2683, [56] := 2683, [57] := 2683, [58] := 2683, [59] := 2683,
        [60] := 2683, [61] := 2683, [62] := 2683, [63] := 2683, [64] := 2683, [65] := 2683, [66] := 2683, [67] := 2683, [68] := 2683, [69] := 2683, [70] := 2683, [71] := 2683, [72] := 2683, [73] := 2683, [74] := 2683, [75] := 2683, [76] := 2683, [77] := 2683, [78] := 2683, [79] := 2683, [80] := 2683, [81] := 2683, [82] := 2683, [83] := 2683, [84] := 2683, [85] := 2683, [86] := 2683, [87] := 2683, [88] := 2683, [89] := 2683, [90] := 2683, [91] := 2683, [92] := 2683, [93] := 2683, [94] := 2683, [95] := 2683, [96] := 2683, [97] := 2683, [98] := 2683, [99] := 2683, [100] := 2683, [101] := 2683, [102] := 2683, [103] := 2683, [104] := 2683, [105] := 2683, [106] := 2683, [107] := 2683, [108] := 2683, [109] := 2683, [110] := 2683, [111] := 2683, [112] := 2683, [113] := 2683, [114] := 2683, [115] := 2683, [116] := 2683, [117] := 2683, [118] := 2683, [119] := 2683,
        [120] := 2683, [121] := 2683, [122] := 2683, [123] := 2683, [124] := 2683, [125] := 2683, [126] := 2683, [127] := 2683, [128] := 2683, [129] := 2683, [130] := 2683, [131] := 2683, [132] := 2683, [133] := 2683, [134] := 2683, [135] := 2683, [136] := 2683, [137] := 2683, [138] := 2683, [139] := 2683, [140] := 2683, [141] := 2683, [142] := 2683, [143] := 2683, [144] := 2683, [145] := 2683, [146] := 2683, [147] := 2683, [148] := 2683, [149] := 2683, [150] := 2683, [151] := 2683, [152] := 2683, [153] := 2683, [154] := 2683, [155] := 2683, [156] := 2683, [157] := 2683, [158] := 2683, [159] := 2683, [160] := 2683, [161] := 2683, [162] := 2683, [163] := 2683, [164] := 2683, [165] := 2683, [166] := 2683, [167] := 2683, [168] := 2683, [169] := 2683, [170] := 2683, [171] := 2683, [172] := 2683, [173] := 2683, [174] := 2683, [175] := 2683, [176] := 2683, [177] := 2683, [178] := 2683, [179] := 2683,
        [180] := 2683, [181] := 2683, [182] := 2683, [183] := 2683, [184] := 2683, [185] := 2683, [186] := 2683, [187] := 2683, [188] := 2683, [189] := 2683, [190] := 2683, [191] := 2683, [192] := 2683, [193] := 2683, [194] := 2683, [195] := 2683, [196] := 2683, [197] := 2683, [198] := 2683, [199] := 2683, [200] := 2683, [201] := 2683, [202] := 2683, [203] := 2683, [204] := 2683, [205] := 2683, [206] := 2683, [207] := 2683, [208] := 2683, [209] := 2683, [210] := 2683, [211] := 2683, [212] := 2683, [213] := 2683, [214] := 2683, [215] := 2683, [216] := 2683, [217] := 2683, [218] := 2683, [219] := 2683, [220] := 2683, [221] := 2683, [222] := 2683, [223] := 2683, [224] := 2683, [225] := 2683, [226] := 2683, [227] := 2683, [228] := 2683, [229] := 2683, [230] := 2683, [231] := 2683, [232] := 2683, [233] := 2683, [234] := 2683, [235] := 2683, [236] := 2683, [237] := 2683, [238] := 2683, [239] := 2683,
        [240] := 2683, [241] := 2683, [242] := 2683, [243] := 2683, [244] := 2683, [245] := 2683, [246] := 2683, [247] := 2683, [248] := 2683, [249] := 2683, [250] := 2683, [251] := 2683, [252] := 2683, [253] := 2683, [254] := 2683, [255] := 2683, [256] := 2683, [257] := 2683, [258] := 2683, [259] := 2683, [260] := 2683, [261] := 2683, [262] := 2683, [263] := 2683, [264] := 2683, [265] := 2683, [266] := 2683, [267] := 2683, [268] := 2683, [269] := 2683, [270] := 2683, [271] := 2683, [272] := 2683, [273] := 2683, [274] := 2683, [275] := 2683, [276] := 2683, [277] := 2683, [278] := 2683, [279] := 2683, [280] := 2683, [281] := 2683, [282] := 2683, [283] := 2683, [284] := 2683, [285] := 2683, [286] := 2683, [287] := 2683, [288] := 2683, [289] := 2683, [290] := 2683, [291] := 2683, [292] := 2683, [293] := 2683, [294] := 2683, [295] := 2683, [296] := 2683, [297] := 2683, [298] := 2683, [299] := 2683,
        [300] := 2683, [301] := 2683, [302] := 2683, [303] := 2686, [304] := 2676, [305] := 2681, [306] := 2679, [307] := 2686, [308] := 2679, [309] := 2691, [310] := 2679, [311] := 2681, [312] := 2681, [313] := 2688, [314] := 2688, [315] := 2686, [316] := 2683, [317] := 2686, [318] := 2693, [319] := 2787, [320] := 2794, [321] := 2787, [322] := 2785, [323] := 2792, [324] := 2794, [325] := 2792, [326] := 2785, [327] := 2783, [328] := 2787, [329] := 2797, [330] := 2792, [331] := 2799, [332] := 2792, [333] := 2818, [334] := 2790, [335] := 2792, [336] := 2783, [337] := 2783, [338] := 2792, [339] := 2794, [340] := 2797, [341] := 2792, [342] := 2794, [343] := 2787, [344] := 2787, [345] := 2783, [346] := 2785, [347] := 2797, [348] := 2794, [349] := 2787, [350] := 2787, [351] := 2780, [352] := 2790, [353] := 2787, [354] := 2794, [355] := 2792, [356] := 2783, [357] := 2787, [358] := 2783, [359] := 2809,
        [360] := 2806, [361] := 2828, [362] := 2813, [363] := 2804, [364] := 2794, [365] := 2790, [366] := 2794, [367] := 2794, [368] := 2790, [369] := 2794, [370] := 2787, [371] := 2797, [372] := 2797, [373] := 2792, [374] := 2799, [375] := 2792, [376] := 2792, [377] := 2787, [378] := 2785, [379] := 2802, [380] := 2799, [381] := 2794, [382] := 2792, [383] := 2794, [384] := 2787, [385] := 2797, [386] := 2797, [387] := 2794, [388] := 2787, [389] := 2794, [390] := 2787, [391] := 2792, [392] := 2790, [393] := 2797, [394] := 2794, [395] := 2794, [396] := 2787, [397] := 2794, [398] := 2787, [399] := 2799, [400] := 2799, [401] := 2797, [402] := 2794, [403] := 2790, [404] := 2787, [405] := 2787, [406] := 2818, [407] := 2811, [408] := 2806, [409] := 2799, [410] := 2790, [411] := 2792, [412] := 2785, [413] := 2787, [414] := 2792, [415] := 2799, [416] := 2802, [417] := 2797, [418] := 2806, [419] := 2802,
        [420] := 2792, [421] := 2799, [422] := 2804, [423] := 2813, [424] := 2792, [425] := 2828, [426] := 2809, [427] := 2783, [428] := 2832, [429] := 2806, [430] := 2811, [431] := 2804, [432] := 2804, [433] := 2813, [434] := 2804, [435] := 2809, [436] := 2816, [437] := 2816, [438] := 2811, [439] := 2811, [440] := 2806, [441] := 2828, [442] := 2792, [443] := 2816, [444] := 2806, [445] := 2797, [446] := 2816, [447] := 2799, [448] := 2799, [449] := 2811, [450] := 2799, [451] := 2797, [452] := 2797, [453] := 2802, [454] := 2778, [455] := 2776, [456] := 2783, [457] := 2792, [458] := 2769, [459] := 2776, [460] := 2776, [461] := 2769, [462] := 2771, [463] := 2769, [464] := 2769, [465] := 2773, [466] := 2769, [467] := 2776, [468] := 2764, [469] := 2766, [470] := 2683, [471] := 2686, [472] := 2702, [473] := 2691, [474] := 2705, [475] := 2688, [476] := 2698, [477] := 2700, [478] := 2686, [479] := 2702,
        [480] := 2683, [481] := 2691, [482] := 2695, [483] := 2688, [484] := 2712, [485] := 2691, [486] := 2700, [487] := 2698, [488] := 2695, [489] := 2700, [490] := 2691, [491] := 2693, [492] := 2693, [493] := 2693, [494] := 2707, [495] := 2695, [496] := 2693, [497] := 2693, [498] := 2683, [499] := 2681, [500] := 2688, [501] := 2691, [502] := 2688, [503] := 2691, [504] := 2681, [505] := 2681, [506] := 2688, [507] := 2686, [508] := 2693, [509] := 2681, [510] := 2676, [511] := 2674, [512] := 2683, [513] := 2693, [514] := 2693, [515] := 2681, [516] := 2683, [517] := 2681, [518] := 2693, [519] := 2688, [520] := 2683, [521] := 2681, [522] := 2676, [523] := 2679, [524] := 2688, [525] := 2693, [526] := 2681, [527] := 2679, [528] := 2679, [529] := 2695, [530] := 2686, [531] := 2679, [532] := 2676, [533] := 2679, [534] := 2688, [535] := 2686, [536] := 2688, [537] := 2679, [538] := 2679, [539] := 2676,
        [540] := 2686, [541] := 2686, [542] := 2676, [543] := 2676, [544] := 2674, [545] := 2681, [546] := 2691, [547] := 2688, [548] := 2688, [549] := 2693, [550] := 2705, [551] := 2681, [552] := 2681, [553] := 2719, [554] := 2688, [555] := 2695, [556] := 2702, [557] := 2688, [558] := 2688, [559] := 2700, [560] := 2700, [561] := 2679, [562] := 2681, [563] := 2688, [564] := 2681, [565] := 2681, [566] := 2686, [567] := 2681, [568] := 2683, [569] := 2693, [570] := 2686, [571] := 2676, [572] := 2679, [573] := 2681, [574] := 2683, [575] := 2686, [576] := 2693, [577] := 2679, [578] := 2679, [579] := 2681, [580] := 2679, [581] := 2688, [582] := 2683, [583] := 2674, [584] := 2681, [585] := 2676, [586] := 2679, [587] := 2681, [588] := 2686, [589] := 2698, [590] := 2683, [591] := 2683, [592] := 2679, [593] := 2686, [594] := 2771, [595] := 2780, [596] := 2780, [597] := 2778, [598] := 2776, [599] := 2773,
        [600] := 2780, [601] := 2771, [602] := 2780, [603] := 2785, [604] := 2778, [605] := 2773, [606] := 2773, [607] := 2783, [608] := 2769, [609] := 2780, [610] := 2780, [611] := 2773, [612] := 2780, [613] := 2771, [614] := 2778, [615] := 2769, [616] := 2769, [617] := 2790, [618] := 2776, [619] := 2783, [620] := 2771, [621] := 2778, [622] := 2773, [623] := 2776, [624] := 2780, [625] := 2773, [626] := 2790, [627] := 2769, [628] := 2785, [629] := 2780, [630] := 2773, [631] := 2787, [632] := 2778, [633] := 2783, [634] := 2776, [635] := 2776, [636] := 2776, [637] := 2783, [638] := 2787, [639] := 2776, [640] := 2783, [641] := 2776, [642] := 2773, [643] := 2783, [644] := 2769, [645] := 2776, [646] := 2776, [647] := 2773, [648] := 2769, [649] := 2778, [650] := 2780, [651] := 2773, [652] := 2783, [653] := 2773, [654] := 2773, [655] := 2773, [656] := 2776, [657] := 2785, [658] := 2778, [659] := 2785,
        [660] := 2771, [661] := 2776, [662] := 2778, [663] := 2776, [664] := 2778, [665] := 2771, [666] := 2787, [667] := 2773, [668] := 2783, [669] := 2787, [670] := 2773, [671] := 2773, [672] := 2771, [673] := 2776, [674] := 2778, [675] := 2790, [676] := 2766, [677] := 2787, [678] := 2785, [679] := 2780, [680] := 2785, [681] := 2771, [682] := 2778, [683] := 2771, [684] := 2780, [685] := 2771, [686] := 2766, [687] := 2776, [688] := 2776, [689] := 2769, [690] := 2773, [691] := 2773, [692] := 2771, [693] := 2776, [694] := 2778, [695] := 2766, [696] := 2771, [697] := 2783, [698] := 2761, [699] := 2766, [700] := 2778, [701] := 2776, [702] := 2776, [703] := 2757, [704] := 2757, [705] := 2759, [706] := 2750, [707] := 2778, [708] := 2776, [709] := 2764, [710] := 2759, [711] := 2757, [712] := 2766, [713] := 2757, [714] := 2757, [715] := 2757, [716] := 2676, [717] := 2683, [718] := 2691, [719] := 2691,
        [720] := 2686, [721] := 2681, [722] := 2688, [723] := 2679, [724] := 2688, [725] := 2691, [726] := 2693, [727] := 2683, [728] := 2681, [729] := 2683, [730] := 2681, [731] := 2693, [732] := 2693, [733] := 2695, [734] := 2698, [735] := 2693, [736] := 2698, [737] := 2693, [738] := 2693, [739] := 2691, [740] := 2702, [741] := 2695, [742] := 2712, [743] := 2693, [744] := 2717, [745] := 2702, [746] := 2709, [747] := 2707, [748] := 2695, [749] := 2679, [750] := 2731, [751] := 2783, [752] := 2794, [753] := 2785, [754] := 2783, [755] := 2794, [756] := 2792, [757] := 2787, [758] := 2787, [759] := 2797, [760] := 2787, [761] := 2785, [762] := 2792, [763] := 2787, [764] := 2787, [765] := 2806, [766] := 2780, [767] := 2783, [768] := 2794, [769] := 2783, [770] := 2783, [771] := 2794, [772] := 2790, [773] := 2783, [774] := 2790, [775] := 2794, [776] := 2785, [777] := 2785, [778] := 2790, [779] := 2792,
        [780] := 2783, [781] := 2790, [782] := 2790, [783] := 2778, [784] := 2787, [785] := 2790, [786] := 2787, [787] := 2783, [788] := 2802, [789] := 2787, [790] := 2794, [791] := 2790, [792] := 2773, [793] := 2776, [794] := 2778, [795] := 2783, [796] := 2776, [797] := 2787, [798] := 2776, [799] := 2787, [800] := 2776, [801] := 2787, [802] := 2769, [803] := 2780, [804] := 2771, [805] := 2787, [806] := 2773, [807] := 2785, [808] := 2771, [809] := 2785, [810] := 2776, [811] := 2778, [812] := 2773, [813] := 2780, [814] := 2771, [815] := 2783, [816] := 2778, [817] := 2780, [818] := 2790, [819] := 2778, [820] := 2785, [821] := 2771, [822] := 2785, [823] := 2776, [824] := 2787, [825] := 2776, [826] := 2787, [827] := 2773, [828] := 2780, [829] := 2773, [830] := 2780, [831] := 2783, [832] := 2785, [833] := 2769, [834] := 2787, [835] := 2766, [836] := 2778, [837] := 2778, [838] := 2776, [839] := 2787,